VERSION : 0.1
   VAR_INPUT
      Enable : Bool;
      CycleTime : Time;
      PulseDuration : Time;
      NowTime : Time;
   END_VAR
   VAR_OUTPUT
      Q_Pulse : Bool;
   END_VAR
   VAR
      CycleTimer : TON;
      PulseTimer : TON;
      State : Int;
      S_PEXT : Int;
   END_VAR
   VAR_TEMP
      PulseActive : Bool;
      StartPulse : Bool;
      TriggerPulse : Bool;
      PulseBusy : Bool;
      DummyWord : Word;
      DummyWord2 : Bool;
      T1 : Int;
      PulseStartTime : Time;
      LastPulseEndTime : Time;
      LastPulseTime : Time;
   END_VAR
BEGIN
   // Logica
   IF #Enable THEN
       // Start cyclische timer
       #CycleTimer(IN := TRUE,
                   PT := #CycleTime);

       IF #CycleTimer.Q THEN
           // Start puls-timer als cyclus voorbij is
           #PulseTimer(IN := TRUE,
                       PT := #PulseDuration);

           // Reset de CycleTimer voor de volgende cyclus
           #CycleTimer(IN := FALSE,
                       PT := #CycleTime);
       END_IF;

       // Puls-timer logica
       IF #PulseTimer.IN THEN
           #Q_Pulse := TRUE;

           IF #PulseTimer.Q THEN
               // Puls voorbij, pulse output uit
               #PulseTimer(IN := FALSE,
                           PT := #PulseDuration);
               #Q_Pulse := FALSE;
           END_IF;
       ELSE
           #Q_Pulse := FALSE;
       END_IF;

   ELSE
       // Alles resetten bij disable
       #CycleTimer(IN := FALSE,
                   PT := #CycleTime);
       #PulseTimer(IN := FALSE,
                   PT := #PulseDuration);
       #Q_Pulse := FALSE;
   END_IF;
END_FUNCTION_BLOCK

FUNCTION_BLOCK "ProductBuffer"   // FB17, SCL
{ S7_Optimized_Access := 'FALSE' }
VERSION : 0.1
   VAR_INPUT
      SensorInput : Bool;
      TimeDelay : Time;
      TriggerFeedback : Bool;
   END_VAR
   VAR_OUTPUT
      TriggerMovement : Bool;
      ProductCount : Int;
   END_VAR
   VAR
      PrevSensor : Bool;
      DelayTimer : TON;
      MovementActive : Bool;
   END_VAR
BEGIN
   // Flankdetectie op sensor
   IF #SensorInput AND NOT #PrevSensor THEN
       IF #ProductCount < 32767 THEN
           #ProductCount := #ProductCount + 1;
       END_IF;
   END_IF;
   #PrevSensor := #SensorInput;

   // Timer mag alleen lopen als:
   // - Er producten zijn
   // - Er geen beweging actief is
   IF (#ProductCount > 0) AND (NOT #MovementActive) THEN
       #DelayTimer(IN := TRUE,
                   PT := #TimeDelay);
   ELSE
       #DelayTimer(IN := FALSE,
                   PT := #TimeDelay);
   END_IF;

   // Als de timer klaar is → activeer beweging en zet MovementActive
   IF #DelayTimer.Q THEN
       #TriggerMovement := TRUE;
       #MovementActive := TRUE;
       #ProductCount := #ProductCount - 1;
       #DelayTimer(IN := FALSE,
                   PT := #TimeDelay); // Reset timer
   END_IF;

   // Wacht op TriggerFeedback om TriggerMovement terug laag te zetten
   IF #MovementActive AND #TriggerFeedback THEN
       #TriggerMovement := FALSE;
       #MovementActive := FALSE;
   END_IF;
END_FUNCTION_BLOCK

FUNCTION_BLOCK "ProductBuffer_V2"   // FB18, SCL
{ S7_Optimized_Access := 'FALSE' }
VERSION : 0.1
   VAR_INPUT
      SensorInput : Bool;
      SensorManual : Bool;
      TimeDelay : Time;
      SystemTime : Time;
      TriggerFeedback : Bool;
   END_VAR
   VAR_OUTPUT
      TriggerMovement : Bool;
      InsertIndex : Int;
      ProductCount : Int;
      SystemTicks : DInt;
   END_VAR
   VAR
      ProductQueue : Array[0..1] of "ProductEntry";
      StartTimes : Struct
         _0 : Time;
         _1 : Time;
         _2 : Time;
         _3 : Time;
         _4 : Time;
         _5 : Time;
         _6 : Time;
         _7 : Time;
         _8 : Time;
         _9 : Time;
      END_STRUCT;
      Actives : Struct
         _0 : Bool;
         _1 : Bool;
         _2 : Bool;
         _3 : Bool;
         _4 : Bool;
         _5 : Bool;
         _6 : Bool;
         _7 : Bool;
         _8 : Bool;
         _9 : Bool;
      END_STRUCT;
      PrevSensor : Bool;
      MovementActive : Bool;
      i : Int;
      Elapsed : DInt;
   END_VAR
BEGIN
   // Flankdetectie sensor
   IF #SensorInput AND NOT #PrevSensor THEN
       CASE #InsertIndex MOD 10 OF
           0:
               IF NOT #Actives._0 THEN
                   #Actives._0 := TRUE;
                   #StartTimes._0 := #SystemTime;
               END_IF;
           1:
               IF NOT #Actives._1 THEN
                   #Actives._1 := TRUE;
                   #StartTimes._1 := #SystemTime;
               END_IF;
           2:
               IF NOT #Actives._2 THEN
                   #Actives._2 := TRUE;
                   #StartTimes._2 := #SystemTime;
               END_IF;
           3:
               IF NOT #Actives._3 THEN
                   #Actives._3 := TRUE;
                   #StartTimes._3 := #SystemTime;
               END_IF;
           4:
               IF NOT #Actives._4 THEN
                   #Actives._4 := TRUE;
                   #StartTimes._4 := #SystemTime;
               END_IF;
           5:
               IF NOT #Actives._5 THEN
                   #Actives._5 := TRUE;
                   #StartTimes._5 := #SystemTime;
               END_IF;
           6:
               IF NOT #Actives._6 THEN
                   #Actives._6 := TRUE;
                   #StartTimes._6 := #SystemTime;
               END_IF;
           7:
               IF NOT #Actives._7 THEN
                   #Actives._7 := TRUE;
                   #StartTimes._7 := #SystemTime;
               END_IF;
           8:
               IF NOT #Actives._8 THEN
                   #Actives._8 := TRUE;
                   #StartTimes._8 := #SystemTime;
               END_IF;
           9:
               IF NOT #Actives._9 THEN
                   #Actives._9 := TRUE;
                   #StartTimes._9 := #SystemTime;
               END_IF;
       END_CASE;
       #InsertIndex := (#InsertIndex + 1) MOD 10;
   END_IF;

   #PrevSensor := #SensorInput;

   // Tellen hoeveel producten actief zijn
   #ProductCount := 0;
   IF #Actives._0 THEN
       #ProductCount := #ProductCount + 1;
   END_IF;
   IF #Actives._1 THEN
       #ProductCount := #ProductCount + 1;
   END_IF;
   IF #Actives._2 THEN
       #ProductCount := #ProductCount + 1;
   END_IF;
   IF #Actives._3 THEN
       #ProductCount := #ProductCount + 1;
   END_IF;
   IF #Actives._4 THEN
       #ProductCount := #ProductCount + 1;
   END_IF;
   IF #Actives._5 THEN
       #ProductCount := #ProductCount + 1;
   END_IF;
   IF #Actives._6 THEN
       #ProductCount := #ProductCount + 1;
   END_IF;
   IF #Actives._7 THEN
       #ProductCount := #ProductCount + 1;
   END_IF;
   IF #Actives._8 THEN
       #ProductCount := #ProductCount + 1;
   END_IF;
   IF #Actives._9 THEN
       #ProductCount := #ProductCount + 1;
   END_IF;

   // Beweging starten als een product klaar is en geen andere beweging actief is
   IF NOT #MovementActive THEN
       IF #Actives._0 THEN
           #Elapsed := TIME_TO_DINT(#SystemTime) - TIME_TO_DINT(#StartTimes._0);
           IF #Elapsed >= TIME_TO_DINT(#TimeDelay) THEN
               #TriggerMovement := TRUE;
               #MovementActive := TRUE;
               #Actives._0 := FALSE;
           END_IF;
       ELSIF #Actives._1 THEN
           #Elapsed := TIME_TO_DINT(#SystemTime) - TIME_TO_DINT(#StartTimes._1);
           IF #Elapsed >= TIME_TO_DINT(#TimeDelay) THEN
               #TriggerMovement := TRUE;
               #MovementActive := TRUE;
               #Actives._1 := FALSE;
           END_IF;
       ELSIF #Actives._2 THEN
           #Elapsed := TIME_TO_DINT(#SystemTime) - TIME_TO_DINT(#StartTimes._2);
           IF #Elapsed >= TIME_TO_DINT(#TimeDelay) THEN
               #TriggerMovement := TRUE;
               #MovementActive := TRUE;
               #Actives._2 := FALSE;
           END_IF;
       ELSIF #Actives._3 THEN
           #Elapsed := TIME_TO_DINT(#SystemTime) - TIME_TO_DINT(#StartTimes._3);
           IF #Elapsed >= TIME_TO_DINT(#TimeDelay) THEN
               #TriggerMovement := TRUE;
               #MovementActive := TRUE;
               #Actives._3 := FALSE;
           END_IF;
       ELSIF #Actives._4 THEN
           #Elapsed := TIME_TO_DINT(#SystemTime) - TIME_TO_DINT(#StartTimes._4);
           IF #Elapsed >= TIME_TO_DINT(#TimeDelay) THEN
               #TriggerMovement := TRUE;
               #MovementActive := TRUE;
               #Actives._4 := FALSE;
           END_IF;
       ELSIF #Actives._5 THEN
           #Elapsed := TIME_TO_DINT(#SystemTime) - TIME_TO_DINT(#StartTimes._5);
           IF #Elapsed >= TIME_TO_DINT(#TimeDelay) THEN
               #TriggerMovement := TRUE;
               #MovementActive := TRUE;
               #Actives._5 := FALSE;
           END_IF;
       ELSIF #Actives._6 THEN
           #Elapsed := TIME_TO_DINT(#SystemTime) - TIME_TO_DINT(#StartTimes._6);
           IF #Elapsed >= TIME_TO_DINT(#TimeDelay) THEN
               #TriggerMovement := TRUE;
               #MovementActive := TRUE;
               #Actives._6 := FALSE;
           END_IF;
       ELSIF #Actives._7 THEN
           #Elapsed := TIME_TO_DINT(#SystemTime) - TIME_TO_DINT(#StartTimes._7);
           IF #Elapsed >= TIME_TO_DINT(#TimeDelay) THEN
               #TriggerMovement := TRUE;
               #MovementActive := TRUE;
               #Actives._7 := FALSE;
           END_IF;
       ELSIF #Actives._8 THEN
           #Elapsed := TIME_TO_DINT(#SystemTime) - TIME_TO_DINT(#StartTimes._8);
           IF #Elapsed >= TIME_TO_DINT(#TimeDelay) THEN
               #TriggerMovement := TRUE;
               #MovementActive := TRUE;
               #Actives._8 := FALSE;
           END_IF;
       ELSIF #Actives._9 THEN
           #Elapsed := TIME_TO_DINT(#SystemTime) - TIME_TO_DINT(#StartTimes._9);
           IF #Elapsed >= TIME_TO_DINT(#TimeDelay) THEN
               #TriggerMovement := TRUE;
               #MovementActive := TRUE;
               #Actives._9 := FALSE;
           END_IF;
       END_IF;
   END_IF;

   // Beweging beëindigen na feedback
   IF #MovementActive AND #TriggerFeedback THEN
       #TriggerMovement := FALSE;
       #MovementActive := FALSE;
   END_IF;
END_FUNCTION_BLOCK

FUNCTION "SCL_Block" : Void   // FC10, SCL
{ S7_Optimized_Access := 'FALSE' }
VERSION : 0.1
BEGIN
   // Reset de Word variabelen aan het begin van elke cyclus
   "Alarms".AlarmsWord := 0;
   "Alarms".HMI_Alarm_Drive1 := 0;
   "Alarms".HMI_Alarm_Drive2 := 0;
   "Alarms".HMI_Alarm_Drive3 := 0;
   "Alarms".HMI_Alarm_Drive4 := 0;
   "Alarms".HMI_Alarm_Drive5 := 0;

   // Controleer de alarmen en zet de respectievelijke bits aan
   IF "Alarms".AlarmStruct.Alarm_Product_Not_Position THEN
       "Alarms".AlarmsWord := "Alarms".AlarmsWord OR WORD#1; // Zet bit 0 aan
   END_IF;

   IF "Alarms".AlarmStruct.Alarm_Axis_Not_Position THEN
       "Alarms".AlarmsWord := "Alarms".AlarmsWord OR WORD#2; // Zet bit 1 aan
   END_IF;

   IF "Alarms".AlarmStruct.Alarm_Drive1 THEN
       "Alarms".HMI_Alarm_Drive1 := "Alarms".HMI_Alarm_Drive1 OR WORD#1; // Zet bit 2 aan
   END_IF;

   IF "Alarms".AlarmStruct.Alarm_Drive2 THEN
       "Alarms".HMI_Alarm_Drive2 := "Alarms".HMI_Alarm_Drive2 OR WORD#1; // Zet bit 3 aan
   END_IF;

   IF "Alarms".AlarmStruct.Alarm_Drive3 THEN
       "Alarms".HMI_Alarm_Drive3 := "Alarms".HMI_Alarm_Drive3 OR WORD#1; // Zet bit 4 aan
   END_IF;

   IF "Alarms".AlarmStruct.Alarm_Drive4 THEN
       "Alarms".HMI_Alarm_Drive4 := "Alarms".HMI_Alarm_Drive4 OR WORD#1; // Zet bit 5 aan
   END_IF;

   IF "Alarms".AlarmStruct.Alarm_Drive5 THEN
       "Alarms".HMI_Alarm_Drive5 := "Alarms".HMI_Alarm_Drive5 OR WORD#1; // Zet bit 6 aan
   END_IF;


   // Position Program Axis 3 (Wals)

   // Configureer de timer om elke 0,5 seconde af te lopen
   "Timer_0_5s".TON(IN := TRUE,
   PT := "PLCMemory"."Encoder PulsOffset");

   // Controleer of de timer is afgelopen
   IF "Timer_0_5s".Q THEN
       // Verhoog of verlaag de positie afhankelijk van de aandrijfsignalen
       IF "Drive 3 RUN FWD" THEN
           "PLCMemory".EncoderPosition := "PLCMemory".EncoderPosition + "PLCMemory".StepSize; // Verhoog met de stepgrootte
       ELSIF "Drive 3 REV" THEN
           "PLCMemory".EncoderPosition := "PLCMemory".EncoderPosition - "PLCMemory".StepSize; // Verlaag met de stepgrootte
       END_IF;

       // Wrapping van de positie bij overschrijden van 360 graden of onder 0 graden
       IF "PLCMemory".EncoderPosition >= 360.0 THEN
           "PLCMemory".EncoderPosition := 0.0;  // Wrapping naar 0 als de positie 360 overschrijdt
       ELSIF "PLCMemory".EncoderPosition < 0.0 THEN
           "PLCMemory".EncoderPosition := 360.0; // Wrapping naar 360 als de positie onder 0 gaat
       END_IF;

       // Reset de timer
       "Timer_0_5s".TON (IN := FALSE,
                         PT := "PLCMemory"."Encoder PulsOffset"); // Reset de timer zodat deze opnieuw kan starten
   END_IF;

   // Homing logica
   IF "Sensor Wals (Option)" THEN
       "PLCMemory".EncoderPosition := 0.0;  // Reset de positie naar 0 als de sensor wordt geactiveerd
   END_IF;



   //Drive Servo Control Here:
   /// Desired Position Axis 3

   // Controleer of de HMI-knop is ingedrukt en er een gewenste positie is ingesteld
   //IF "HMI_Des_Pos_Axis3" THEN
       //"GoButtonPressed" := TRUE; // HMI-knop is ingedrukt, start beweging
   //END_IF;

   // Beveiliging voor de Desired_Encoder_Position: Zorg dat de waarde tussen 0 en 360 blijft
   //IF "PLCMemory".Desired_Encoder_Position > 360.0 THEN
     //  "PLCMemory".Desired_Encoder_Position := 360.0;  // Zet naar 360 als de waarde boven 360 ligt
   //ELSIF "PLCMemory".Desired_Encoder_Position < 0.0 THEN
       //"PLCMemory".Desired_Encoder_Position := 0.0;  // Zet naar 0 als de waarde onder 0 ligt
   //END_IF;

   // Wrapping van de gewenste positie: Als de gewenste positie 360 is, zet deze dan op 0
   //IF "PLCMemory".Desired_Encoder_Position = 360.0 THEN
      // "PLCMemory".Desired_Encoder_Position := 0.0;  // Wrapping naar 0 als de gewenste positie 360 is
   //END_IF;

   // Voer beweging uit totdat de gewenste positie is bereikt
   //IF "GoButtonPressed" THEN
       // Bepaal de bewegingsrichting en start de beweging
     //  IF "PLCMemory".EncoderPosition < "PLCMemory".Desired_Encoder_Position - "PLCMemory".Tolerance THEN
           // Beweeg vooruit met StepSize als snelheid
         //  "PLCMemory".EncoderPosition := "PLCMemory".EncoderPosition + "PLCMemory".StepSize;
        //   "Drive_3_Manual" := TRUE;   // Activeer vooruitbeweging
         //  "Drive 3 REV" := FALSE;     // Zorg dat achteruitbeweging uit is

     //  ELSIF "PLCMemory".EncoderPosition > "PLCMemory".Desired_Encoder_Position + "PLCMemory".Tolerance THEN
           // Beweeg achteruit met StepSize als snelheid
        //   "PLCMemory".EncoderPosition := "PLCMemory".EncoderPosition - "PLCMemory".StepSize;
       //    "Drive_3_Manual" := FALSE;  // Zorg dat vooruitbeweging uit is
       //    "Drive 3 REV" := TRUE;      // Activeer achteruitbeweging

      // ELSE
           // Stop de beweging zodra de positie binnen de tolerantie komt
         //  "Drive_3_Manual" := FALSE;    // Zet vooruitbeweging uit
        //   "Drive 3 REV" := FALSE;       // Zet achteruitbeweging uit
        //   "GoButtonPressed" := FALSE;   // Zet de Go-knop uit om verdere beweging te stoppen
      // END_IF;
   //END_IF;
END_FUNCTION

FUNCTION "SafetyFunction_Block" : Void   // FC12, LAD
{ S7_Optimized_Access := 'FALSE' }
VERSION : 0.1
   VAR_INPUT
      "ESB NC Contact" : Bool;
      "ESB NO Contact" : Bool;
      "Reset NO Contact" : Bool;
      "SAFE door 1 NC Contact" : Bool;
      "SAFE door 2 NC Contact" : Bool;
      "Safety Relais NO Contact" : Bool;
   END_VAR
   VAR_OUTPUT
      SAFE_OK_Signal : Bool;
   END_VAR
BEGIN

REGION Network 1: +MC-21K6:1 - Noodstop Circuit
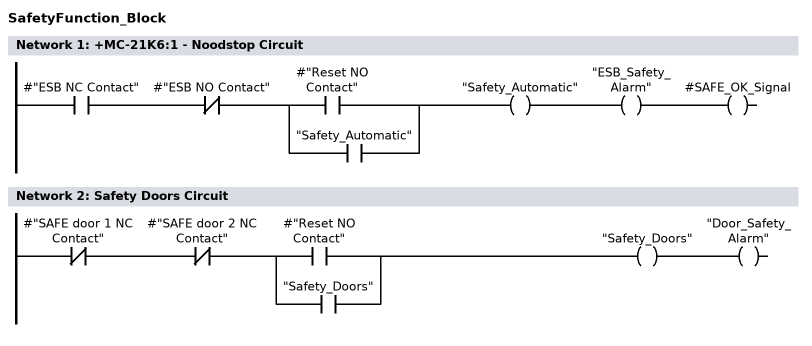
   RUNG wire#powerrail
      Contact( #"ESB NC Contact" )
      I_Contact( #"ESB NO Contact" )
      wire#w1
      Contact( #"Reset NO Contact" )
      wire#w2
      Coil( "Safety_Automatic" )
      Coil( "ESB_Safety_Alarm" )
      Coil( #SAFE_OK_Signal )
   END_RUNG
   RUNG wire#w1
      Contact( "Safety_Automatic" )
   END_RUNG wire#w2
   // the same network as SCL:
   "Safety_Automatic" := #"ESB NC Contact" AND NOT #"ESB NO Contact" AND (#"Reset NO Contact" OR "Safety_Automatic");
   "ESB_Safety_Alarm" := "Safety_Automatic";
   #SAFE_OK_Signal := "Safety_Automatic";
END_REGION

REGION Network 2: Safety Doors Circuit
   RUNG wire#powerrail
      I_Contact( #"SAFE door 1 NC Contact" )
      I_Contact( #"SAFE door 2 NC Contact" )
      wire#w1
      Contact( #"Reset NO Contact" )
      wire#w2
      Coil( "Safety_Doors" )
      Coil( "Door_Safety_Alarm" )
   END_RUNG
   RUNG wire#w1
      Contact( "Safety_Doors" )
   END_RUNG wire#w2
   // the same network as SCL:
   "Safety_Doors" := NOT #"SAFE door 1 NC Contact" AND NOT #"SAFE door 2 NC Contact" AND (#"Reset NO Contact" OR "Safety_Doors");
   "Door_Safety_Alarm" := "Safety_Doors";
END_REGION
END_FUNCTION

FUNCTION "SystemRUN_Block" : Void   // FC13, LAD
{ S7_Optimized_Access := 'FALSE' }
VERSION : 0.1
   VAR_INPUT
      "Safety Relais Contact" : Bool;
      "Stop Machine NC Contact" : Bool;
      "Fill Magzine Contact" : Bool;
      "Start Machine NO Contact" : Bool;
   END_VAR
   VAR_OUTPUT
      "Run Output Lamp" : Bool;
   END_VAR
BEGIN

REGION Network 1: Systeem RUN
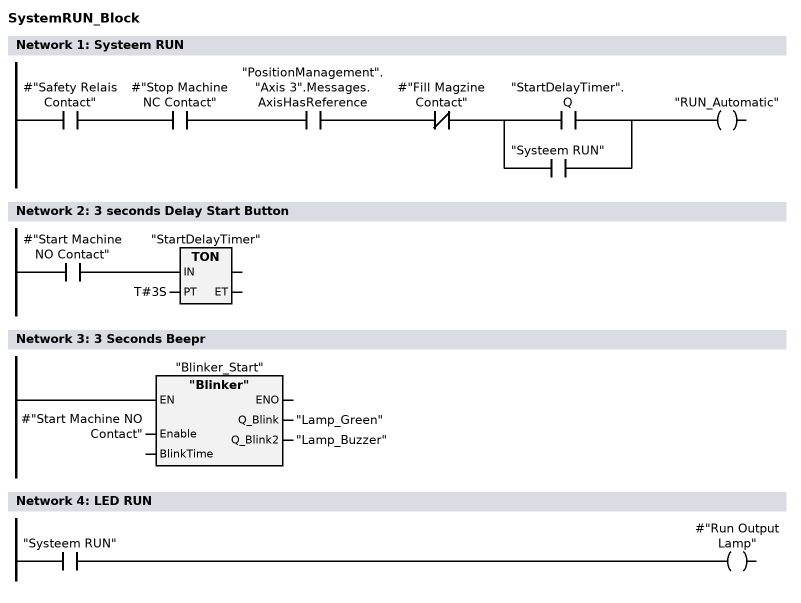
   RUNG wire#powerrail
      Contact( #"Safety Relais Contact" )
      Contact( #"Stop Machine NC Contact" )
      Contact( "PositionManagement"."Axis 3".Messages.AxisHasReference )
      I_Contact( #"Fill Magzine Contact" )
      wire#w1
      Contact( "StartDelayTimer".Q )
      wire#w2
      Coil( "RUN_Automatic" )
   END_RUNG
   RUNG wire#w1
      Contact( "Systeem RUN" )
   END_RUNG wire#w2
   // the same network as SCL:
   "RUN_Automatic" := #"Safety Relais Contact" AND #"Stop Machine NC Contact" AND "PositionManagement"."Axis 3".Messages.AxisHasReference AND NOT #"Fill Magzine Contact" AND ("StartDelayTimer".Q OR "Systeem RUN");
END_REGION

REGION Network 2: 3 seconds Delay Start Button
   "StartDelayTimer".TON(IN := #"Start Machine NO Contact", PT := T#3S);
END_REGION

REGION Network 3: 3 Seconds Beepr
   RUNG wire#powerrail
      "Blinker_Start"(Enable := #"Start Machine NO Contact", BlinkTime :=, Q_Blink => "Lamp_Green", Q_Blink2 => "Lamp_Buzzer")
   END_RUNG
   // the same network as SCL:
   "Blinker_Start"(Enable := #"Start Machine NO Contact", Q_Blink => "Lamp_Green", Q_Blink2 => "Lamp_Buzzer");   // "Blinker"
END_REGION

REGION Network 4: LED RUN
   RUNG wire#powerrail
      Contact( "Systeem RUN" )
      Coil( #"Run Output Lamp" )
   END_RUNG
   // the same network as SCL:
   #"Run Output Lamp" := "Systeem RUN";
END_REGION
END_FUNCTION

FUNCTION "SiemensEnc" : Void   // FC15, STL
TITLE = Test Siemens ENCODER
{ S7_Optimized_Access := 'FALSE' }
VERSION : 0.1
BEGIN

REGION Network 1: Presettings
         L     0;  //Delete control bits
         T     %DB1.DBD0;
         T     %DB1.DBD4;
         SET;
         S     %DB1.DBX4.0;  //Open SW gate
END_REGION

REGION Network 2: Write to the control interface
END_REGION

REGION Network 3: Read from the feedback interface
   //Read 8 bytes from the 1 Count24V
   //Configured start address of inputs
         L     "Tag_25":P;
         T     %DB1.DBD8;
         L     "Tag_26":P;
         T     %DB1.DBD12;
         R     %DB1.DBX4.0;  //Close SW gate
END_REGION
END_FUNCTION

// folder: Motion

FUNCTION_BLOCK "MC_Move"   // FB10, FBD
TITLE = MC_Move
{ S7_Optimized_Access := 'FALSE' }
VERSION : 0.1
// Block moves an Axis to an Desired Position, this block comes with the brake feature. When the axis is on position it keeps the brake for a time. You can set the time in the Brake Time field.
   VAR_INPUT
      Start : Bool;
      "Desired Position" : Real;
      "Speed (50-75%)" : Int;
      "Brake on Position" : Bool;
      Acceleration : Real;
      Deacceleration : Real;
      "Drive Ready" : Bool;
      "Drive On Position" : Bool;
      "Brake Time" : Time := T#500ms;
      "Safety OK" : Bool;
   END_VAR
   VAR_OUTPUT
      Go : Bool;
      "Desired Position Out" : Real;
      "Speed Output" : Int;
      "Acceleration Out" : Real;
      "Deacceleration Out" : Real;
      "Brake Out" : Bool;
   END_VAR
   VAR_TEMP
      SR_1 : Bool;
   END_VAR
BEGIN

REGION Network 1: Start - Go To Position + Speed
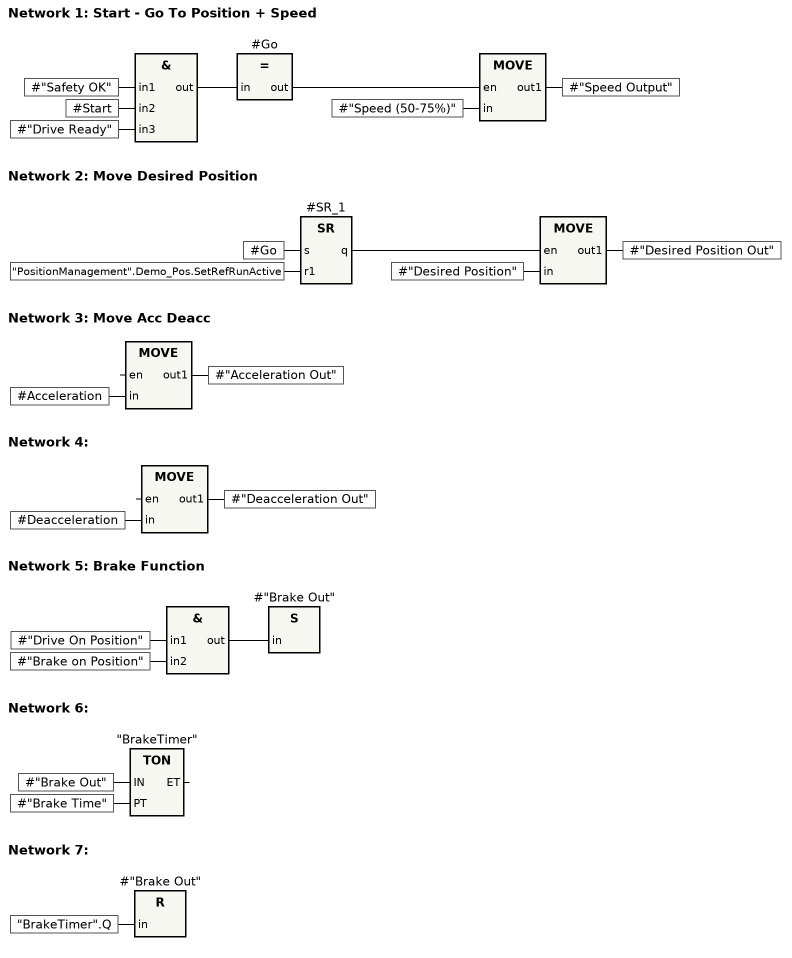
   #Go := #"Safety OK" AND #Start AND #"Drive Ready";
   IF #Go THEN #"Speed Output" := #"Speed (50-75%)"; END_IF;
END_REGION

REGION Network 2: Move Desired Position
   IF #Go THEN
       #SR_1 := TRUE;   // SR flip-flop
   END_IF;
   IF "PositionManagement".Demo_Pos.SetRefRunActive THEN #SR_1 := FALSE; END_IF;
   IF #SR_1 THEN #"Desired Position Out" := #"Desired Position"; END_IF;
END_REGION

REGION Network 3: Move Acc Deacc
   #"Acceleration Out" := #Acceleration;
END_REGION

REGION Network 4
   #"Deacceleration Out" := #Deacceleration;
END_REGION

REGION Network 5: Brake Function
   IF #"Drive On Position" AND #"Brake on Position" THEN #"Brake Out" := TRUE; END_IF;
END_REGION

REGION Network 6
   "BrakeTimer".TON(IN := #"Brake Out", PT := #"Brake Time");
END_REGION

REGION Network 7
   IF "BrakeTimer".Q THEN #"Brake Out" := FALSE; END_IF;
END_REGION
END_FUNCTION_BLOCK

FUNCTION_BLOCK "MC_Jog"   // FB11, FBD
TITLE = MC_Jog
{ S7_Optimized_Access := 'FALSE' }
VERSION : 0.1
// With this block you can Jog an Axis manual, you can set the speed on 25%, 50% or 75%. It also has an brake functionality, when you set Brake to true, it holds the brake for 2 seconds, then releases it.
   VAR_INPUT
      "Jog Forward" : Bool;
      "Jog Backward" : Bool;
      Speed : Int;
      Brake : Bool;
   END_VAR
   VAR_OUTPUT
      "Drive Fwd Output" : Bool;
      "Drive Rev Output" : Bool;
      "Drive Speed Output" : Int;
      "Drive Brake Output" : Bool;
   END_VAR
BEGIN

REGION Network 1: Manual Control
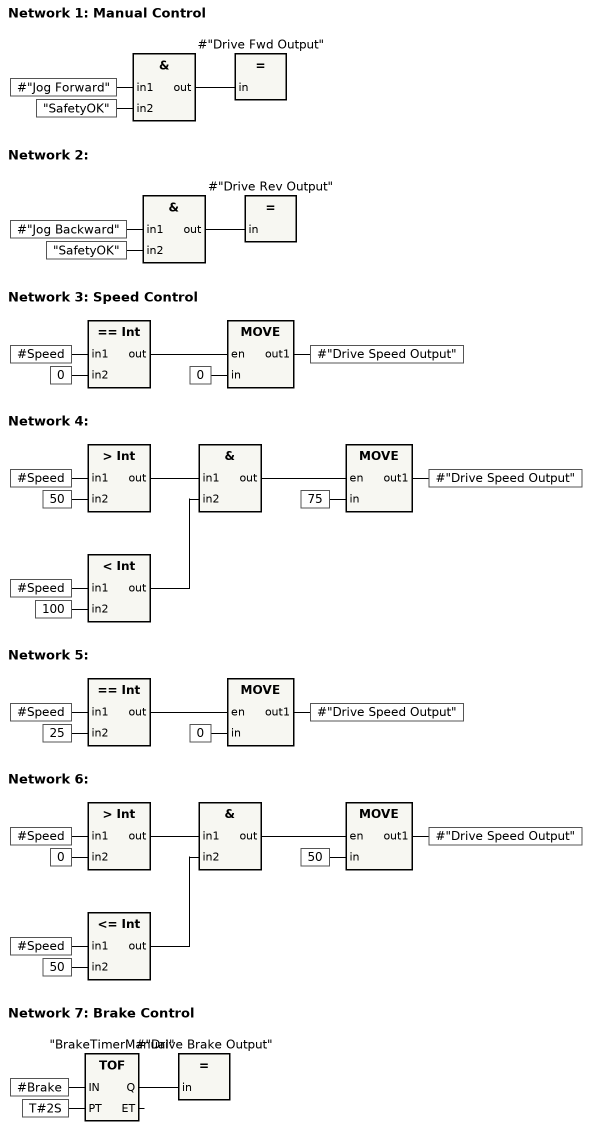
   #"Drive Fwd Output" := #"Jog Forward" AND "SafetyOK";
END_REGION

REGION Network 2
   #"Drive Rev Output" := #"Jog Backward" AND "SafetyOK";
END_REGION

REGION Network 3: Speed Control
   IF #Speed = 0 THEN #"Drive Speed Output" := 0; END_IF;
END_REGION

REGION Network 4
   IF (#Speed > 50) AND (#Speed < 100) THEN #"Drive Speed Output" := 75; END_IF;
END_REGION

REGION Network 5
   IF #Speed = 25 THEN #"Drive Speed Output" := 0; END_IF;
END_REGION

REGION Network 6
   IF (#Speed > 0) AND (#Speed <= 50) THEN #"Drive Speed Output" := 50; END_IF;
END_REGION

REGION Network 7: Brake Control
   "BrakeTimerManual".TOF(IN := #Brake, PT := T#2S);
   #"Drive Brake Output" := "BrakeTimerManual".Q;
END_REGION
END_FUNCTION_BLOCK

FUNCTION "Axis_Confirmation" : Void   // FC7, FBD
TITLE = Axis Confirmation Block
{ S7_Optimized_Access := 'FALSE' }
VERSION : 0.1
   VAR_INPUT
      "Set Position" : Real;
   END_VAR
   VAR_OUTPUT
      "Axis On Position" : Bool;
      Min_Position_1 : Real;
      Max_Position_1 : Real;
   END_VAR
BEGIN

REGION Network 2: Calculate Position Tolerance 1
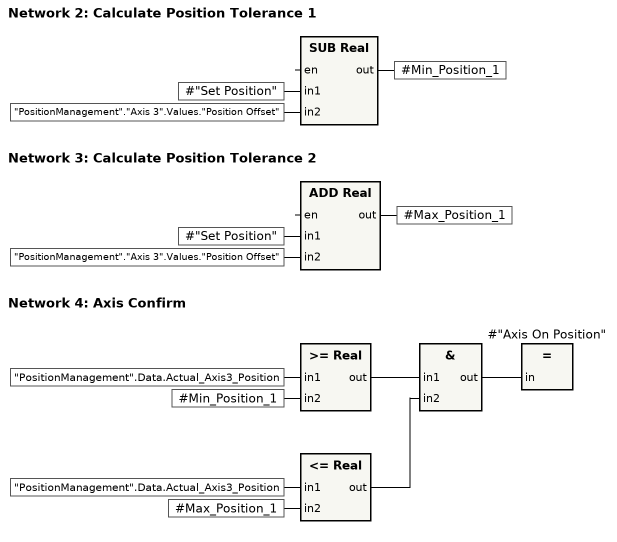
   #Min_Position_1 := #"Set Position" - "PositionManagement"."Axis 3".Values."Position Offset";
END_REGION

REGION Network 3: Calculate Position Tolerance 2
   #Max_Position_1 := #"Set Position" + "PositionManagement"."Axis 3".Values."Position Offset";
END_REGION

REGION Network 4: Axis Confirm
   #"Axis On Position" := ("PositionManagement".Data.Actual_Axis3_Position >= #Min_Position_1) AND ("PositionManagement".Data.Actual_Axis3_Position <= #Max_Position_1);
END_REGION
END_FUNCTION

FUNCTION "EMStopDrives_Block" : Void   // FC14, LAD
{ S7_Optimized_Access := 'FALSE' }
VERSION : 0.1
   VAR_INPUT
      "Safety Callback" : Bool;
      Direct_Stop : Bool;
   END_VAR
   VAR_OUTPUT
      "Drive 1 Brake Out" : Bool;
      "Drive 2 Brake Out" : Bool;
      "Drive 3 Brake Out" : Bool;
      "Drive 4 Brake Out" : Bool;
      "Drive 5 Brake Out" : Bool;
      "Drive 6 Brake Out" : Bool;
      "Drive 7 Brake Out" : Bool;
      "Drive 8 Brake Out" : Bool;
      "Drive 9 Brake Out" : Bool;
      "Drive 10 Brake Out" : Bool;
   END_VAR
BEGIN

REGION Network 1: Drives Emergency Stop
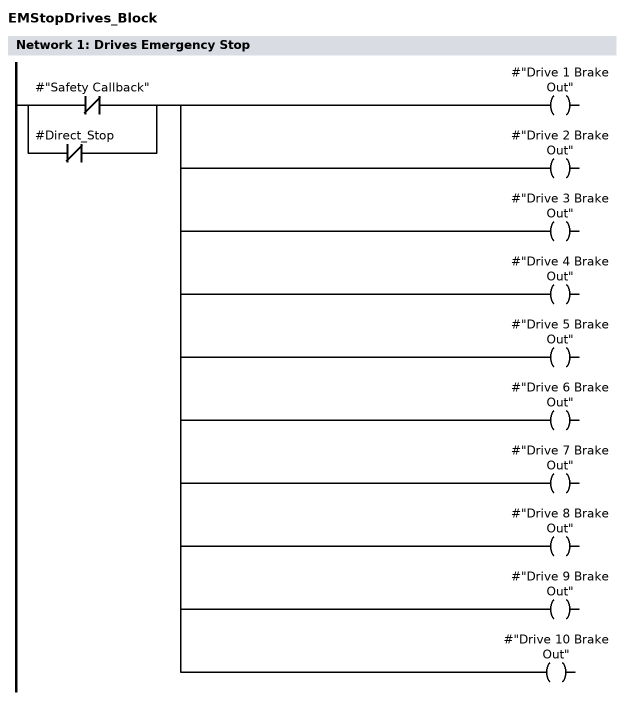
   RUNG wire#powerrail
      I_Contact( #"Safety Callback" )
      wire#w1
      Coil( #"Drive 1 Brake Out" )
   END_RUNG
   RUNG wire#powerrail
      I_Contact( #Direct_Stop )
   END_RUNG wire#w1
   RUNG wire#w1
      Coil( #"Drive 2 Brake Out" )
   END_RUNG
   RUNG wire#w1
      Coil( #"Drive 3 Brake Out" )
   END_RUNG
   RUNG wire#w1
      Coil( #"Drive 4 Brake Out" )
   END_RUNG
   RUNG wire#w1
      Coil( #"Drive 5 Brake Out" )
   END_RUNG
   RUNG wire#w1
      Coil( #"Drive 6 Brake Out" )
   END_RUNG
   RUNG wire#w1
      Coil( #"Drive 7 Brake Out" )
   END_RUNG
   RUNG wire#w1
      Coil( #"Drive 8 Brake Out" )
   END_RUNG
   RUNG wire#w1
      Coil( #"Drive 9 Brake Out" )
   END_RUNG
   RUNG wire#w1
      Coil( #"Drive 10 Brake Out" )
   END_RUNG
   // the same network as SCL:
   #"Drive 1 Brake Out" := NOT #"Safety Callback" OR NOT #Direct_Stop;
   #"Drive 2 Brake Out" := #"Drive 1 Brake Out";
   #"Drive 3 Brake Out" := #"Drive 1 Brake Out";
   #"Drive 4 Brake Out" := #"Drive 1 Brake Out";
   #"Drive 5 Brake Out" := #"Drive 1 Brake Out";
   #"Drive 6 Brake Out" := #"Drive 1 Brake Out";
   #"Drive 7 Brake Out" := #"Drive 1 Brake Out";
   #"Drive 8 Brake Out" := #"Drive 1 Brake Out";
   #"Drive 9 Brake Out" := #"Drive 1 Brake Out";
   #"Drive 10 Brake Out" := #"Drive 1 Brake Out";
END_REGION
END_FUNCTION

FUNCTION "EncoderFeedback" : Void   // FC16, FBD
TITLE = EncoderFeedback Block
{ S7_Optimized_Access := 'FALSE' }
VERSION : 0.1
   VAR_INPUT
      CounterTag : Int;   // Connect to the CounterTag IW102
      Position_Offset : Real;   // Fill in the tolerance, when the axis approves the position. Above or below the desired position
      Pulsfactor : Real;   // Number of pulses after 360 degree turn of the axis.
      Position_Correction : Real;   // Small Position Correction for the Axis
      ReferenceRun_Command : Bool;   // Command of starting the referencerun
      ReferenceSwitch : Bool;   // ReferenceSwitch Mounted on Axis
      ReferencePosition : Int;   // Position where the index puls of the reference switch enters.
   END_VAR
   VAR_OUTPUT
      Scaled_Position : Real;   // Scaled Position scaled with Pulsfactor
      Actual_Enc_Pos : Real;   // Actual Encoder Position
      AxisDB_Connection : Real;   // Connection with Axis DB connection
   END_VAR
   VAR_TEMP
      Corrected_Axis_Pos : Real;
      Unscaled_Position : Int;   // Unscaled Position of the Encoder
      Unsc2 : Int;   // Unsc 2 position
      Act_Enc_Pos_Int : DInt;
      Scaled_Position_Real : Real;
      PosDint : DInt;
      Unscaled_Position_Real : Real;
      InternalCounter : Int;
      CalDifCounter : Int;
      Pos_Storage : Int;
      Pos_Diffrence : Int;
      Add_Pos : Int;
      Sub_Pos : Int;
      LessThanZero : Bool;
      LTZ_out : Int;
   END_VAR
BEGIN

REGION Network 1: SPARE
END_REGION

REGION Network 2 (STL): Call the Countermodule
         L     #CounterTag;  //Van tellerkaart TAG Gelinkt aan IW102
         L     "PositionManagement".Data.CntPlsPrev;  //Vorige scan
         -D;
         T     "PositionManagement".Data.CntPlsDiff;  //Verschil

         L     "PositionManagement".Data.CntPlsDiff;  // Verschil groter dan nul?
         L     0;
         >D;
         JCN   chkneg;

         L     "PositionManagement".Data.CntPlsDiff;  //Verschil optellen bij actuele pulswaarde
         L     "PositionManagement".Data.CntPlsAct;
         +D;
         T     "PositionManagement".Data.CntPlsAct;
         JU    end;  //rest overslaan.

   chkneg:L     "PositionManagement".Data.CntPlsDiff;  // Verschil groter dan nul?
         L     0;
         <D;
         JCN   end;
         L     -1;  //verschil positief maken
         *D;
         T     "PositionManagement".Data.CntPlsDiff;  //verschil positief

         L     "PositionManagement".Data.CntPlsAct;  //Verschil optellen bij actuele pulswaarde
         +D;
         T     "PositionManagement".Data.CntPlsAct;

   end:  NOP   0;

         L     #CounterTag;
         T     "PositionManagement".Data.CntPlsPrev;
END_REGION

REGION Network 3: Store Old Position
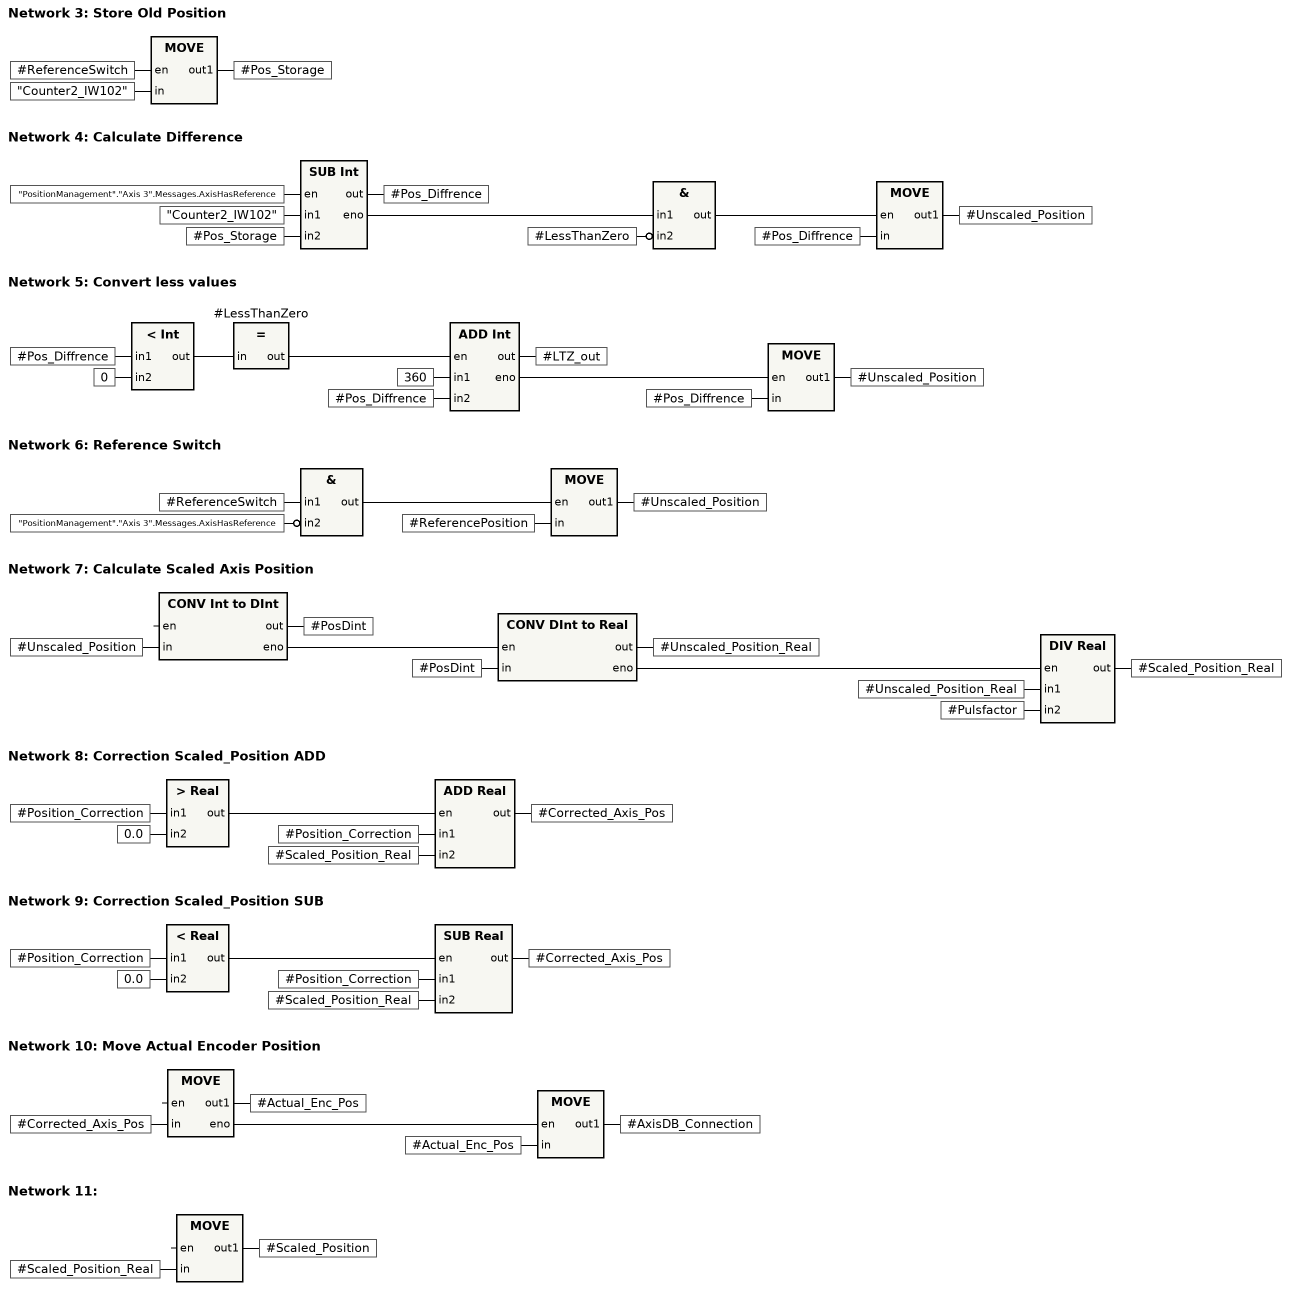
   IF #ReferenceSwitch THEN #Pos_Storage := "Counter2_IW102"; END_IF;
END_REGION

REGION Network 4: Calculate Difference
   // ENO of a box is taken as its EN; it also drops when the box reports an error
   IF "PositionManagement"."Axis 3".Messages.AxisHasReference THEN
       #Pos_Diffrence := "Counter2_IW102" - #Pos_Storage;
   END_IF;
   IF "PositionManagement"."Axis 3".Messages.AxisHasReference AND NOT #LessThanZero THEN
       #Unscaled_Position := #Pos_Diffrence;
   END_IF;
END_REGION

REGION Network 5: Convert less values
   // ENO of a box is taken as its EN; it also drops when the box reports an error
   #LessThanZero := #Pos_Diffrence < 0;
   IF #LessThanZero THEN
       #LTZ_out := 360 + #Pos_Diffrence;
       #Unscaled_Position := #Pos_Diffrence;
   END_IF;
END_REGION

REGION Network 6: Reference Switch
   IF #ReferenceSwitch AND NOT "PositionManagement"."Axis 3".Messages.AxisHasReference THEN
       #Unscaled_Position := #ReferencePosition;
   END_IF;
END_REGION

REGION Network 7: Calculate Scaled Axis Position
   // ENO of a box is taken as its EN; it also drops when the box reports an error
   #PosDint := INT_TO_DINT(#Unscaled_Position);
   #Unscaled_Position_Real := DINT_TO_REAL(#PosDint);
   #Scaled_Position_Real := #Unscaled_Position_Real / #Pulsfactor;
END_REGION

REGION Network 8: Correction Scaled_Position ADD
   IF #Position_Correction > 0.0 THEN
       #Corrected_Axis_Pos := #Position_Correction + #Scaled_Position_Real;
   END_IF;
END_REGION

REGION Network 9: Correction Scaled_Position SUB
   IF #Position_Correction < 0.0 THEN
       #Corrected_Axis_Pos := #Position_Correction - #Scaled_Position_Real;
   END_IF;
END_REGION

REGION Network 10: Move Actual Encoder Position
   // ENO of a box is taken as its EN; it also drops when the box reports an error
   #Actual_Enc_Pos := #Corrected_Axis_Pos;
   #AxisDB_Connection := #Actual_Enc_Pos;
END_REGION

REGION Network 11
   #Scaled_Position := #Scaled_Position_Real;
END_REGION
END_FUNCTION

FUNCTION "Servo_DriveManager" : Void   // FC17, FBD
TITLE = Drive Manager Closed Loop
{ S7_Optimized_Access := 'FALSE' }
VERSION : 0.1
// Drive Manager for Closed Loop with Encoder
   VAR_INPUT
      "[NAME] Axis Name" : String;
      "[INPUT] ReferenceSwitch_Input" : Bool;
      "[INPUT] Drive Ready" : Bool;
      "[INPUT] E-STOP Check" : Bool;
      "[COMMAND] Start_Reference Run" : Bool;
      "[COMMAND] Take_over_Pos" : Bool;
      "[COMMAND] Go to Position" : Bool;
      "[COMMAND] Axis Manual Forward" : Bool;
      "[COMMAND] Axis Manual Reverse" : Bool;
      "[COMMAND] Axis Speed" : Int;
      "[COMMAND] Axis Fast Stop" : Bool;
      "[COMMAND] Go To Rest" : Bool;
      "[COMMAND] Axis Brake" : Bool;
      "[VALUE] Reference Position" : Int;
      "[VALUE] Set Position" : Real;
      "[VALUE] Rest Position" : Real;
      "[VALUE] Accelerating" : Real;
      "[VALUE] Deaccelerating" : Real;
      "[VALUE] Position Tolerance" : Real;
      "[COMMUNICATION] MasterWord" : String;
      "[COMMUNICATION] Callback" : String;
   END_VAR
   VAR_OUTPUT
      "[OUTPUT] Drive FWD Command" : Bool;
      "[OUTPUT] Drive REV Command" : Bool;
      "[OUTPUT] Drive Speed 2 (50%)" : Bool;
      "[OUTPUT] Drive Speed 3 (75%)" : Bool;
      "[OUTPUT] Drive Fast Stop Command" : Bool;
      "[MESSAGE] Axis Busy" : Bool;
      "[MESSAGE] Error Executing" : Bool;
      "[MESSAGE] Axis On Position" : Bool;
      "[MESSAGE] Axis On Rest" : Bool;
      "[MESSAGE] Drive State" : String;
      "[MESSAGE] Axis Slips" : String;
   END_VAR
   VAR_TEMP
      UnscPos : Int;
      ScPos : Real;
      ActEncPos : Real;
      SetRefRun : Bool;
      SetRefRun_Q : Bool;
      MoveToRest : Bool;
      MoveToRest_Q : Bool;
      Automatic_Positive : Bool;
      Manual_Positive : Bool;
      Automatic_Negative : Bool;
      Manual_Negative : Bool;
      HS_Positive : Bool;
      MasterWordHex : Int;
      Speed50 : Bool;
      Speed75 : Bool;
      Min_Position : Real;
      Max_Position : Real;
      Axis_On_Position : Bool;
      Direction_Forward : Bool;
      Direction_Backward : Bool;
      Drive_Auto_Fwd : Bool;
      InternalFastStop : Bool;
      RefRunSetSignal : Bool;
      GoToRest2 : Bool;
      "[COMMAND] Go to Position_Rest" : Bool;
      RestPos_SpareMove : Real;
   END_VAR
   VAR_TEMP   // added for the SCL form of the ladder/FBD networks
      _w1 : Bool;
   END_VAR
BEGIN

REGION Network 1: Reference Run